REGION Network 14: EM - UnSuspending State Complete
   RUNG wire#powerrail
      Contact( "EM01".PackML_Sts.Alarm.sts_UnSuspending_SC )
      wire#w1
      Contact( "EM01".PackML_Sts.CM01.sts_UnSuspending_SC )
      wire#w2
      Contact( "EM01".PackML_Sts.CM02.sts_UnSuspending_SC )
      wire#w3
      Contact( "EM01".PackML_Sts.CM03.sts_UnSuspending_SC )
      wire#w4
      Contact( "EM01".PackML_Sts.CM04.sts_UnSuspending_SC )
      wire#w5
      Contact( "EM01".PackML_Sts.CM05.sts_UnSuspending_SC )
      wire#w6
      Contact( "EM01".PackML_Sts.CM06.sts_UnSuspending_SC )
      wire#w7
      Contact( "EM01".PackML_Sts.CM07.sts_UnSuspending_SC )
      wire#w8
      Contact( "EM01".PackML_Sts.CM08.sts_UnSuspending_SC )
      wire#w9
      Contact( "EM01".PackML_Sts.CM09.sts_UnSuspending_SC )
      wire#w10
      Contact( "EM01".PackML_Sts.CM10.sts_UnSuspending_SC )
      wire#w11
      Coil( "EM01".PackML_Sts.Unit.sts_UnSuspending_SC )
   END_RUNG
   RUNG wire#powerrail
      I_Contact( "EM01".PackML_Sts.Alarm.moduleActive )
   END_RUNG wire#w1
   RUNG wire#w1
      I_Contact( "EM01".PackML_Sts.CM01.moduleActive )
   END_RUNG wire#w2
   RUNG wire#w2
      I_Contact( "EM01".PackML_Sts.CM02.moduleActive )
   END_RUNG wire#w3
   RUNG wire#w3
      I_Contact( "EM01".PackML_Sts.CM03.moduleActive )
   END_RUNG wire#w4
   RUNG wire#w4
      I_Contact( "EM01".PackML_Sts.CM04.moduleActive )
   END_RUNG wire#w5
   RUNG wire#w5
      I_Contact( "EM01".PackML_Sts.CM05.moduleActive )
   END_RUNG wire#w6
   RUNG wire#w6
      I_Contact( "EM01".PackML_Sts.CM06.moduleActive )
   END_RUNG wire#w7
   RUNG wire#w7
      I_Contact( "EM01".PackML_Sts.CM07.moduleActive )
   END_RUNG wire#w8
   RUNG wire#w8
      I_Contact( "EM01".PackML_Sts.CM08.moduleActive )
   END_RUNG wire#w9
   RUNG wire#w9
      I_Contact( "EM01".PackML_Sts.CM09.moduleActive )
   END_RUNG wire#w10
   RUNG wire#w10
      I_Contact( "EM01".PackML_Sts.CM10.moduleActive )
   END_RUNG wire#w11
   // the same network as SCL:
   "EM01".PackML_Sts.Unit.sts_UnSuspending_SC := ("EM01".PackML_Sts.Alarm.sts_UnSuspending_SC OR NOT "EM01".PackML_Sts.Alarm.moduleActive) AND ("EM01".PackML_Sts.CM01.sts_UnSuspending_SC OR NOT "EM01".PackML_Sts.CM01.moduleActive) AND ("EM01".PackML_Sts.CM02.sts_UnSuspending_SC OR NOT "EM01".PackML_Sts.CM02.moduleActive) AND ("EM01".PackML_Sts.CM03.sts_UnSuspending_SC OR NOT "EM01".PackML_Sts.CM03.moduleActive) AND ("EM01".PackML_Sts.CM04.sts_UnSuspending_SC OR NOT "EM01".PackML_Sts.CM04.moduleActive) AND ("EM01".PackML_Sts.CM05.sts_UnSuspending_SC OR NOT "EM01".PackML_Sts.CM05.moduleActive) AND ("EM01".PackML_Sts.CM06.sts_UnSuspending_SC OR NOT "EM01".PackML_Sts.CM06.moduleActive) AND ("EM01".PackML_Sts.CM07.sts_UnSuspending_SC OR NOT "EM01".PackML_Sts.CM07.moduleActive) AND ("EM01".PackML_Sts.CM08.sts_UnSuspending_SC OR NOT "EM01".PackML_Sts.CM08.moduleActive) AND ("EM01".PackML_Sts.CM09.sts_UnSuspending_SC OR NOT "EM01".PackML_Sts.CM09.moduleActive) AND ("EM01".PackML_Sts.CM10.sts_UnSuspending_SC OR NOT "EM01".PackML_Sts.CM10.moduleActive);
END_REGION

REGION Network 15: EM - Abort Command
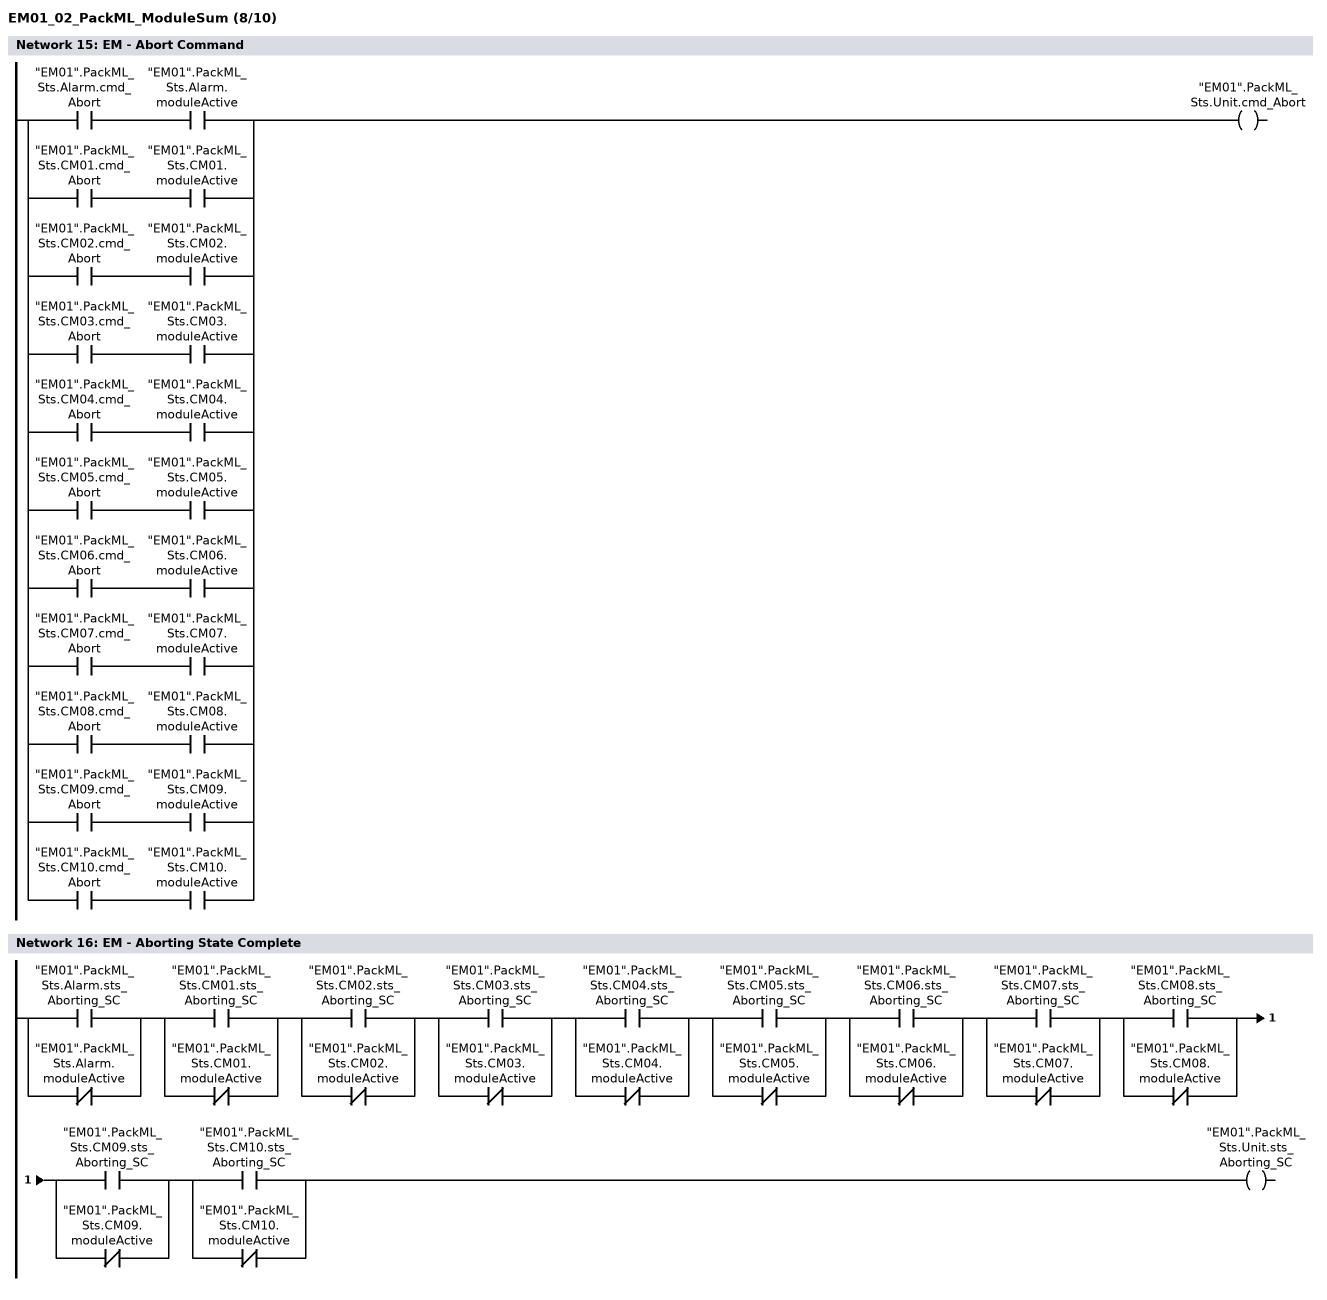
   RUNG wire#powerrail
      Contact( "EM01".PackML_Sts.Alarm.cmd_Abort )
      Contact( "EM01".PackML_Sts.Alarm.moduleActive )
      wire#w1
      Coil( "EM01".PackML_Sts.Unit.cmd_Abort )
   END_RUNG
   RUNG wire#powerrail
      Contact( "EM01".PackML_Sts.CM01.cmd_Abort )
      Contact( "EM01".PackML_Sts.CM01.moduleActive )
   END_RUNG wire#w1
   RUNG wire#powerrail
      Contact( "EM01".PackML_Sts.CM02.cmd_Abort )
      Contact( "EM01".PackML_Sts.CM02.moduleActive )
   END_RUNG wire#w1
   RUNG wire#powerrail
      Contact( "EM01".PackML_Sts.CM03.cmd_Abort )
      Contact( "EM01".PackML_Sts.CM03.moduleActive )
   END_RUNG wire#w1
   RUNG wire#powerrail
      Contact( "EM01".PackML_Sts.CM04.cmd_Abort )
      Contact( "EM01".PackML_Sts.CM04.moduleActive )
   END_RUNG wire#w1
   RUNG wire#powerrail
      Contact( "EM01".PackML_Sts.CM05.cmd_Abort )
      Contact( "EM01".PackML_Sts.CM05.moduleActive )
   END_RUNG wire#w1
   RUNG wire#powerrail
      Contact( "EM01".PackML_Sts.CM06.cmd_Abort )
      Contact( "EM01".PackML_Sts.CM06.moduleActive )
   END_RUNG wire#w1
   RUNG wire#powerrail
      Contact( "EM01".PackML_Sts.CM07.cmd_Abort )
      Contact( "EM01".PackML_Sts.CM07.moduleActive )
   END_RUNG wire#w1
   RUNG wire#powerrail
      Contact( "EM01".PackML_Sts.CM08.cmd_Abort )
      Contact( "EM01".PackML_Sts.CM08.moduleActive )
   END_RUNG wire#w1
   RUNG wire#powerrail
      Contact( "EM01".PackML_Sts.CM09.cmd_Abort )
      Contact( "EM01".PackML_Sts.CM09.moduleActive )
   END_RUNG wire#w1
   RUNG wire#powerrail
      Contact( "EM01".PackML_Sts.CM10.cmd_Abort )
      Contact( "EM01".PackML_Sts.CM10.moduleActive )
   END_RUNG wire#w1
   // the same network as SCL:
   "EM01".PackML_Sts.Unit.cmd_Abort := ("EM01".PackML_Sts.Alarm.cmd_Abort AND "EM01".PackML_Sts.Alarm.moduleActive) OR ("EM01".PackML_Sts.CM01.cmd_Abort AND "EM01".PackML_Sts.CM01.moduleActive) OR ("EM01".PackML_Sts.CM02.cmd_Abort AND "EM01".PackML_Sts.CM02.moduleActive) OR ("EM01".PackML_Sts.CM03.cmd_Abort AND "EM01".PackML_Sts.CM03.moduleActive) OR ("EM01".PackML_Sts.CM04.cmd_Abort AND "EM01".PackML_Sts.CM04.moduleActive) OR ("EM01".PackML_Sts.CM05.cmd_Abort AND "EM01".PackML_Sts.CM05.moduleActive) OR ("EM01".PackML_Sts.CM06.cmd_Abort AND "EM01".PackML_Sts.CM06.moduleActive) OR ("EM01".PackML_Sts.CM07.cmd_Abort AND "EM01".PackML_Sts.CM07.moduleActive) OR ("EM01".PackML_Sts.CM08.cmd_Abort AND "EM01".PackML_Sts.CM08.moduleActive) OR ("EM01".PackML_Sts.CM09.cmd_Abort AND "EM01".PackML_Sts.CM09.moduleActive) OR ("EM01".PackML_Sts.CM10.cmd_Abort AND "EM01".PackML_Sts.CM10.moduleActive);
END_REGION

REGION Network 16: EM - Aborting State Complete
   RUNG wire#powerrail
      Contact( "EM01".PackML_Sts.Alarm.sts_Aborting_SC )
      wire#w1
      Contact( "EM01".PackML_Sts.CM01.sts_Aborting_SC )
      wire#w2
      Contact( "EM01".PackML_Sts.CM02.sts_Aborting_SC )
      wire#w3
      Contact( "EM01".PackML_Sts.CM03.sts_Aborting_SC )
      wire#w4
      Contact( "EM01".PackML_Sts.CM04.sts_Aborting_SC )
      wire#w5
      Contact( "EM01".PackML_Sts.CM05.sts_Aborting_SC )
      wire#w6
      Contact( "EM01".PackML_Sts.CM06.sts_Aborting_SC )
      wire#w7
      Contact( "EM01".PackML_Sts.CM07.sts_Aborting_SC )
      wire#w8
      Contact( "EM01".PackML_Sts.CM08.sts_Aborting_SC )
      wire#w9
      Contact( "EM01".PackML_Sts.CM09.sts_Aborting_SC )
      wire#w10
      Contact( "EM01".PackML_Sts.CM10.sts_Aborting_SC )
      wire#w11
      Coil( "EM01".PackML_Sts.Unit.sts_Aborting_SC )
   END_RUNG
   RUNG wire#powerrail
      I_Contact( "EM01".PackML_Sts.Alarm.moduleActive )
   END_RUNG wire#w1
   RUNG wire#w1
      I_Contact( "EM01".PackML_Sts.CM01.moduleActive )
   END_RUNG wire#w2
   RUNG wire#w2
      I_Contact( "EM01".PackML_Sts.CM02.moduleActive )
   END_RUNG wire#w3
   RUNG wire#w3
      I_Contact( "EM01".PackML_Sts.CM03.moduleActive )
   END_RUNG wire#w4
   RUNG wire#w4
      I_Contact( "EM01".PackML_Sts.CM04.moduleActive )
   END_RUNG wire#w5
   RUNG wire#w5
      I_Contact( "EM01".PackML_Sts.CM05.moduleActive )
   END_RUNG wire#w6
   RUNG wire#w6
      I_Contact( "EM01".PackML_Sts.CM06.moduleActive )
   END_RUNG wire#w7
   RUNG wire#w7
      I_Contact( "EM01".PackML_Sts.CM07.moduleActive )
   END_RUNG wire#w8
   RUNG wire#w8
      I_Contact( "EM01".PackML_Sts.CM08.moduleActive )
   END_RUNG wire#w9
   RUNG wire#w9
      I_Contact( "EM01".PackML_Sts.CM09.moduleActive )
   END_RUNG wire#w10
   RUNG wire#w10
      I_Contact( "EM01".PackML_Sts.CM10.moduleActive )
   END_RUNG wire#w11
   // the same network as SCL:
   "EM01".PackML_Sts.Unit.sts_Aborting_SC := ("EM01".PackML_Sts.Alarm.sts_Aborting_SC OR NOT "EM01".PackML_Sts.Alarm.moduleActive) AND ("EM01".PackML_Sts.CM01.sts_Aborting_SC OR NOT "EM01".PackML_Sts.CM01.moduleActive) AND ("EM01".PackML_Sts.CM02.sts_Aborting_SC OR NOT "EM01".PackML_Sts.CM02.moduleActive) AND ("EM01".PackML_Sts.CM03.sts_Aborting_SC OR NOT "EM01".PackML_Sts.CM03.moduleActive) AND ("EM01".PackML_Sts.CM04.sts_Aborting_SC OR NOT "EM01".PackML_Sts.CM04.moduleActive) AND ("EM01".PackML_Sts.CM05.sts_Aborting_SC OR NOT "EM01".PackML_Sts.CM05.moduleActive) AND ("EM01".PackML_Sts.CM06.sts_Aborting_SC OR NOT "EM01".PackML_Sts.CM06.moduleActive) AND ("EM01".PackML_Sts.CM07.sts_Aborting_SC OR NOT "EM01".PackML_Sts.CM07.moduleActive) AND ("EM01".PackML_Sts.CM08.sts_Aborting_SC OR NOT "EM01".PackML_Sts.CM08.moduleActive) AND ("EM01".PackML_Sts.CM09.sts_Aborting_SC OR NOT "EM01".PackML_Sts.CM09.moduleActive) AND ("EM01".PackML_Sts.CM10.sts_Aborting_SC OR NOT "EM01".PackML_Sts.CM10.moduleActive);
END_REGION

REGION Network 17: EM - Clear Command
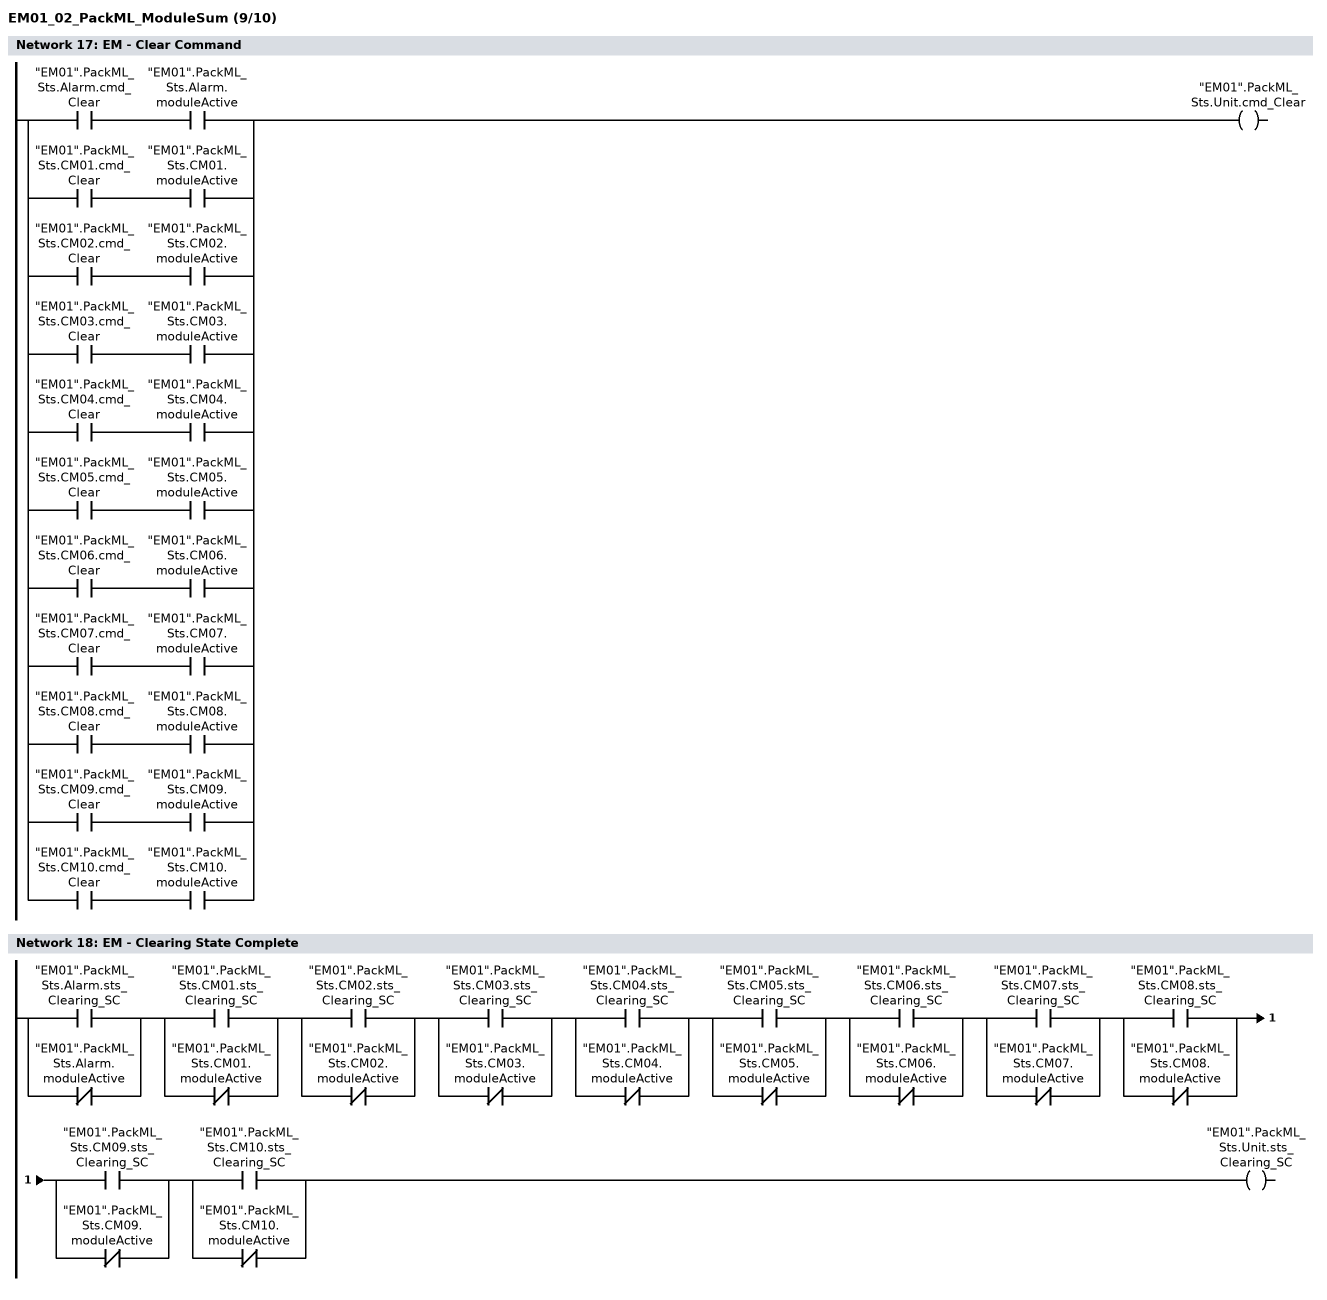
   RUNG wire#powerrail
      Contact( "EM01".PackML_Sts.Alarm.cmd_Clear )
      Contact( "EM01".PackML_Sts.Alarm.moduleActive )
      wire#w1
      Coil( "EM01".PackML_Sts.Unit.cmd_Clear )
   END_RUNG
   RUNG wire#powerrail
      Contact( "EM01".PackML_Sts.CM01.cmd_Clear )
      Contact( "EM01".PackML_Sts.CM01.moduleActive )
   END_RUNG wire#w1
   RUNG wire#powerrail
      Contact( "EM01".PackML_Sts.CM02.cmd_Clear )
      Contact( "EM01".PackML_Sts.CM02.moduleActive )
   END_RUNG wire#w1
   RUNG wire#powerrail
      Contact( "EM01".PackML_Sts.CM03.cmd_Clear )
      Contact( "EM01".PackML_Sts.CM03.moduleActive )
   END_RUNG wire#w1
   RUNG wire#powerrail
      Contact( "EM01".PackML_Sts.CM04.cmd_Clear )
      Contact( "EM01".PackML_Sts.CM04.moduleActive )
   END_RUNG wire#w1
   RUNG wire#powerrail
      Contact( "EM01".PackML_Sts.CM05.cmd_Clear )
      Contact( "EM01".PackML_Sts.CM05.moduleActive )
   END_RUNG wire#w1
   RUNG wire#powerrail
      Contact( "EM01".PackML_Sts.CM06.cmd_Clear )
      Contact( "EM01".PackML_Sts.CM06.moduleActive )
   END_RUNG wire#w1
   RUNG wire#powerrail
      Contact( "EM01".PackML_Sts.CM07.cmd_Clear )
      Contact( "EM01".PackML_Sts.CM07.moduleActive )
   END_RUNG wire#w1
   RUNG wire#powerrail
      Contact( "EM01".PackML_Sts.CM08.cmd_Clear )
      Contact( "EM01".PackML_Sts.CM08.moduleActive )
   END_RUNG wire#w1
   RUNG wire#powerrail
      Contact( "EM01".PackML_Sts.CM09.cmd_Clear )
      Contact( "EM01".PackML_Sts.CM09.moduleActive )
   END_RUNG wire#w1
   RUNG wire#powerrail
      Contact( "EM01".PackML_Sts.CM10.cmd_Clear )
      Contact( "EM01".PackML_Sts.CM10.moduleActive )
   END_RUNG wire#w1
   // the same network as SCL:
   "EM01".PackML_Sts.Unit.cmd_Clear := ("EM01".PackML_Sts.Alarm.cmd_Clear AND "EM01".PackML_Sts.Alarm.moduleActive) OR ("EM01".PackML_Sts.CM01.cmd_Clear AND "EM01".PackML_Sts.CM01.moduleActive) OR ("EM01".PackML_Sts.CM02.cmd_Clear AND "EM01".PackML_Sts.CM02.moduleActive) OR ("EM01".PackML_Sts.CM03.cmd_Clear AND "EM01".PackML_Sts.CM03.moduleActive) OR ("EM01".PackML_Sts.CM04.cmd_Clear AND "EM01".PackML_Sts.CM04.moduleActive) OR ("EM01".PackML_Sts.CM05.cmd_Clear AND "EM01".PackML_Sts.CM05.moduleActive) OR ("EM01".PackML_Sts.CM06.cmd_Clear AND "EM01".PackML_Sts.CM06.moduleActive) OR ("EM01".PackML_Sts.CM07.cmd_Clear AND "EM01".PackML_Sts.CM07.moduleActive) OR ("EM01".PackML_Sts.CM08.cmd_Clear AND "EM01".PackML_Sts.CM08.moduleActive) OR ("EM01".PackML_Sts.CM09.cmd_Clear AND "EM01".PackML_Sts.CM09.moduleActive) OR ("EM01".PackML_Sts.CM10.cmd_Clear AND "EM01".PackML_Sts.CM10.moduleActive);
END_REGION

REGION Network 18: EM - Clearing State Complete
   RUNG wire#powerrail
      Contact( "EM01".PackML_Sts.Alarm.sts_Clearing_SC )
      wire#w1
      Contact( "EM01".PackML_Sts.CM01.sts_Clearing_SC )
      wire#w2
      Contact( "EM01".PackML_Sts.CM02.sts_Clearing_SC )
      wire#w3
      Contact( "EM01".PackML_Sts.CM03.sts_Clearing_SC )
      wire#w4
      Contact( "EM01".PackML_Sts.CM04.sts_Clearing_SC )
      wire#w5
      Contact( "EM01".PackML_Sts.CM05.sts_Clearing_SC )
      wire#w6
      Contact( "EM01".PackML_Sts.CM06.sts_Clearing_SC )
      wire#w7
      Contact( "EM01".PackML_Sts.CM07.sts_Clearing_SC )
      wire#w8
      Contact( "EM01".PackML_Sts.CM08.sts_Clearing_SC )
      wire#w9
      Contact( "EM01".PackML_Sts.CM09.sts_Clearing_SC )
      wire#w10
      Contact( "EM01".PackML_Sts.CM10.sts_Clearing_SC )
      wire#w11
      Coil( "EM01".PackML_Sts.Unit.sts_Clearing_SC )
   END_RUNG
   RUNG wire#powerrail
      I_Contact( "EM01".PackML_Sts.Alarm.moduleActive )
   END_RUNG wire#w1
   RUNG wire#w1
      I_Contact( "EM01".PackML_Sts.CM01.moduleActive )
   END_RUNG wire#w2
   RUNG wire#w2
      I_Contact( "EM01".PackML_Sts.CM02.moduleActive )
   END_RUNG wire#w3
   RUNG wire#w3
      I_Contact( "EM01".PackML_Sts.CM03.moduleActive )
   END_RUNG wire#w4
   RUNG wire#w4
      I_Contact( "EM01".PackML_Sts.CM04.moduleActive )
   END_RUNG wire#w5
   RUNG wire#w5
      I_Contact( "EM01".PackML_Sts.CM05.moduleActive )
   END_RUNG wire#w6
   RUNG wire#w6
      I_Contact( "EM01".PackML_Sts.CM06.moduleActive )
   END_RUNG wire#w7
   RUNG wire#w7
      I_Contact( "EM01".PackML_Sts.CM07.moduleActive )
   END_RUNG wire#w8
   RUNG wire#w8
      I_Contact( "EM01".PackML_Sts.CM08.moduleActive )
   END_RUNG wire#w9
   RUNG wire#w9
      I_Contact( "EM01".PackML_Sts.CM09.moduleActive )
   END_RUNG wire#w10
   RUNG wire#w10
      I_Contact( "EM01".PackML_Sts.CM10.moduleActive )
   END_RUNG wire#w11
   // the same network as SCL:
   "EM01".PackML_Sts.Unit.sts_Clearing_SC := ("EM01".PackML_Sts.Alarm.sts_Clearing_SC OR NOT "EM01".PackML_Sts.Alarm.moduleActive) AND ("EM01".PackML_Sts.CM01.sts_Clearing_SC OR NOT "EM01".PackML_Sts.CM01.moduleActive) AND ("EM01".PackML_Sts.CM02.sts_Clearing_SC OR NOT "EM01".PackML_Sts.CM02.moduleActive) AND ("EM01".PackML_Sts.CM03.sts_Clearing_SC OR NOT "EM01".PackML_Sts.CM03.moduleActive) AND ("EM01".PackML_Sts.CM04.sts_Clearing_SC OR NOT "EM01".PackML_Sts.CM04.moduleActive) AND ("EM01".PackML_Sts.CM05.sts_Clearing_SC OR NOT "EM01".PackML_Sts.CM05.moduleActive) AND ("EM01".PackML_Sts.CM06.sts_Clearing_SC OR NOT "EM01".PackML_Sts.CM06.moduleActive) AND ("EM01".PackML_Sts.CM07.sts_Clearing_SC OR NOT "EM01".PackML_Sts.CM07.moduleActive) AND ("EM01".PackML_Sts.CM08.sts_Clearing_SC OR NOT "EM01".PackML_Sts.CM08.moduleActive) AND ("EM01".PackML_Sts.CM09.sts_Clearing_SC OR NOT "EM01".PackML_Sts.CM09.moduleActive) AND ("EM01".PackML_Sts.CM10.sts_Clearing_SC OR NOT "EM01".PackML_Sts.CM10.moduleActive);
END_REGION

REGION Network 19: EM - Execute State Complete
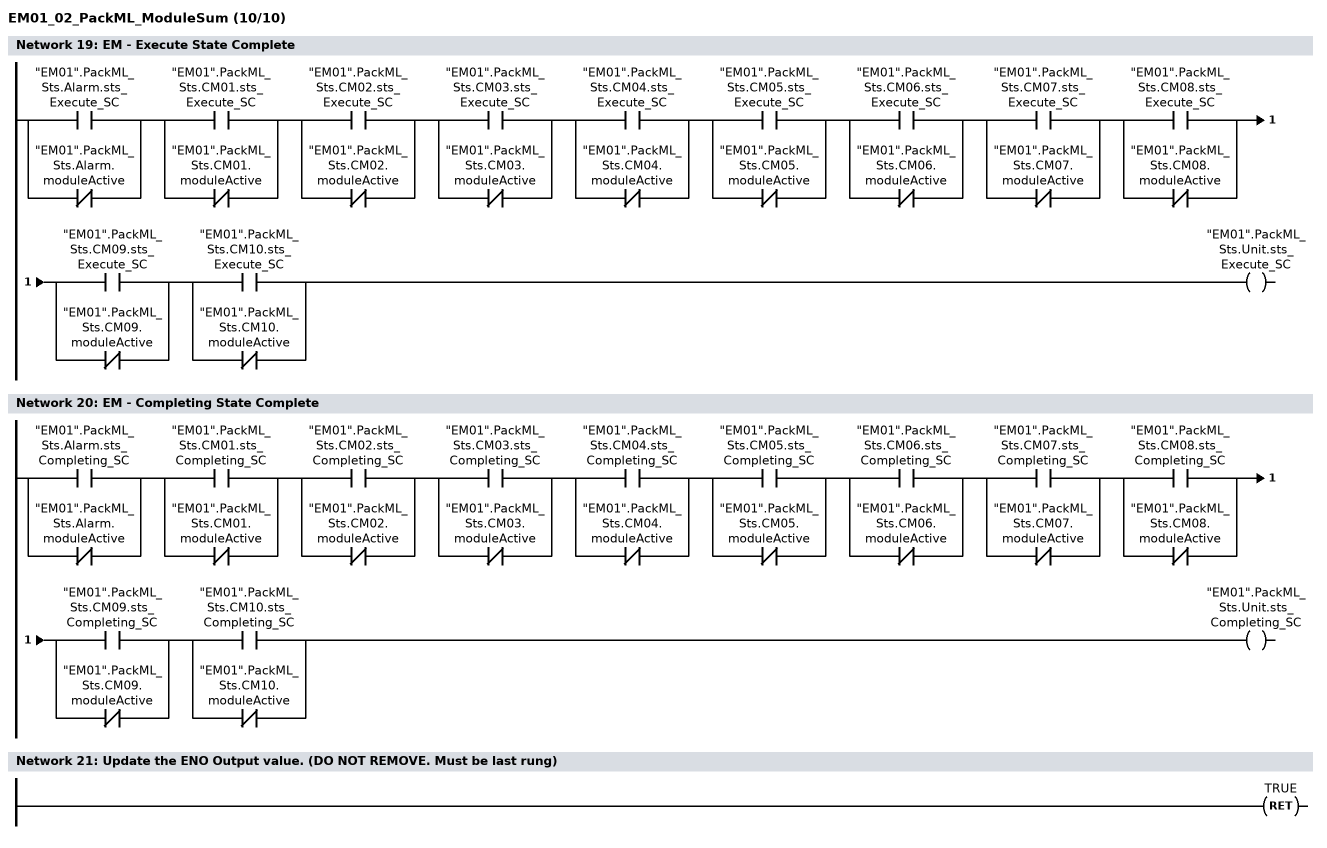
   RUNG wire#powerrail
      Contact( "EM01".PackML_Sts.Alarm.sts_Execute_SC )
      wire#w1
      Contact( "EM01".PackML_Sts.CM01.sts_Execute_SC )
      wire#w2
      Contact( "EM01".PackML_Sts.CM02.sts_Execute_SC )
      wire#w3
      Contact( "EM01".PackML_Sts.CM03.sts_Execute_SC )
      wire#w4
      Contact( "EM01".PackML_Sts.CM04.sts_Execute_SC )
      wire#w5
      Contact( "EM01".PackML_Sts.CM05.sts_Execute_SC )
      wire#w6
      Contact( "EM01".PackML_Sts.CM06.sts_Execute_SC )
      wire#w7
      Contact( "EM01".PackML_Sts.CM07.sts_Execute_SC )
      wire#w8
      Contact( "EM01".PackML_Sts.CM08.sts_Execute_SC )
      wire#w9
      Contact( "EM01".PackML_Sts.CM09.sts_Execute_SC )
      wire#w10
      Contact( "EM01".PackML_Sts.CM10.sts_Execute_SC )
      wire#w11
      Coil( "EM01".PackML_Sts.Unit.sts_Execute_SC )
   END_RUNG
   RUNG wire#powerrail
      I_Contact( "EM01".PackML_Sts.Alarm.moduleActive )
   END_RUNG wire#w1
   RUNG wire#w1
      I_Contact( "EM01".PackML_Sts.CM01.moduleActive )
   END_RUNG wire#w2
   RUNG wire#w2
      I_Contact( "EM01".PackML_Sts.CM02.moduleActive )
   END_RUNG wire#w3
   RUNG wire#w3
      I_Contact( "EM01".PackML_Sts.CM03.moduleActive )
   END_RUNG wire#w4
   RUNG wire#w4
      I_Contact( "EM01".PackML_Sts.CM04.moduleActive )
   END_RUNG wire#w5
   RUNG wire#w5
      I_Contact( "EM01".PackML_Sts.CM05.moduleActive )
   END_RUNG wire#w6
   RUNG wire#w6
      I_Contact( "EM01".PackML_Sts.CM06.moduleActive )
   END_RUNG wire#w7
   RUNG wire#w7
      I_Contact( "EM01".PackML_Sts.CM07.moduleActive )
   END_RUNG wire#w8
   RUNG wire#w8
      I_Contact( "EM01".PackML_Sts.CM08.moduleActive )
   END_RUNG wire#w9
   RUNG wire#w9
      I_Contact( "EM01".PackML_Sts.CM09.moduleActive )
   END_RUNG wire#w10
   RUNG wire#w10
      I_Contact( "EM01".PackML_Sts.CM10.moduleActive )
   END_RUNG wire#w11
   // the same network as SCL:
   "EM01".PackML_Sts.Unit.sts_Execute_SC := ("EM01".PackML_Sts.Alarm.sts_Execute_SC OR NOT "EM01".PackML_Sts.Alarm.moduleActive) AND ("EM01".PackML_Sts.CM01.sts_Execute_SC OR NOT "EM01".PackML_Sts.CM01.moduleActive) AND ("EM01".PackML_Sts.CM02.sts_Execute_SC OR NOT "EM01".PackML_Sts.CM02.moduleActive) AND ("EM01".PackML_Sts.CM03.sts_Execute_SC OR NOT "EM01".PackML_Sts.CM03.moduleActive) AND ("EM01".PackML_Sts.CM04.sts_Execute_SC OR NOT "EM01".PackML_Sts.CM04.moduleActive) AND ("EM01".PackML_Sts.CM05.sts_Execute_SC OR NOT "EM01".PackML_Sts.CM05.moduleActive) AND ("EM01".PackML_Sts.CM06.sts_Execute_SC OR NOT "EM01".PackML_Sts.CM06.moduleActive) AND ("EM01".PackML_Sts.CM07.sts_Execute_SC OR NOT "EM01".PackML_Sts.CM07.moduleActive) AND ("EM01".PackML_Sts.CM08.sts_Execute_SC OR NOT "EM01".PackML_Sts.CM08.moduleActive) AND ("EM01".PackML_Sts.CM09.sts_Execute_SC OR NOT "EM01".PackML_Sts.CM09.moduleActive) AND ("EM01".PackML_Sts.CM10.sts_Execute_SC OR NOT "EM01".PackML_Sts.CM10.moduleActive);
END_REGION

REGION Network 20: EM - Completing State Complete
   RUNG wire#powerrail
      Contact( "EM01".PackML_Sts.Alarm.sts_Completing_SC )
      wire#w1
      Contact( "EM01".PackML_Sts.CM01.sts_Completing_SC )
      wire#w2
      Contact( "EM01".PackML_Sts.CM02.sts_Completing_SC )
      wire#w3
      Contact( "EM01".PackML_Sts.CM03.sts_Completing_SC )
      wire#w4
      Contact( "EM01".PackML_Sts.CM04.sts_Completing_SC )
      wire#w5
      Contact( "EM01".PackML_Sts.CM05.sts_Completing_SC )
      wire#w6
      Contact( "EM01".PackML_Sts.CM06.sts_Completing_SC )
      wire#w7
      Contact( "EM01".PackML_Sts.CM07.sts_Completing_SC )
      wire#w8
      Contact( "EM01".PackML_Sts.CM08.sts_Completing_SC )
      wire#w9
      Contact( "EM01".PackML_Sts.CM09.sts_Completing_SC )
      wire#w10
      Contact( "EM01".PackML_Sts.CM10.sts_Completing_SC )
      wire#w11
      Coil( "EM01".PackML_Sts.Unit.sts_Completing_SC )
   END_RUNG
   RUNG wire#powerrail
      I_Contact( "EM01".PackML_Sts.Alarm.moduleActive )
   END_RUNG wire#w1
   RUNG wire#w1
      I_Contact( "EM01".PackML_Sts.CM01.moduleActive )
   END_RUNG wire#w2
   RUNG wire#w2
      I_Contact( "EM01".PackML_Sts.CM02.moduleActive )
   END_RUNG wire#w3
   RUNG wire#w3
      I_Contact( "EM01".PackML_Sts.CM03.moduleActive )
   END_RUNG wire#w4
   RUNG wire#w4
      I_Contact( "EM01".PackML_Sts.CM04.moduleActive )
   END_RUNG wire#w5
   RUNG wire#w5
      I_Contact( "EM01".PackML_Sts.CM05.moduleActive )
   END_RUNG wire#w6
   RUNG wire#w6
      I_Contact( "EM01".PackML_Sts.CM06.moduleActive )
   END_RUNG wire#w7
   RUNG wire#w7
      I_Contact( "EM01".PackML_Sts.CM07.moduleActive )
   END_RUNG wire#w8
   RUNG wire#w8
      I_Contact( "EM01".PackML_Sts.CM08.moduleActive )
   END_RUNG wire#w9
   RUNG wire#w9
      I_Contact( "EM01".PackML_Sts.CM09.moduleActive )
   END_RUNG wire#w10
   RUNG wire#w10
      I_Contact( "EM01".PackML_Sts.CM10.moduleActive )
   END_RUNG wire#w11
   // the same network as SCL:
   "EM01".PackML_Sts.Unit.sts_Completing_SC := ("EM01".PackML_Sts.Alarm.sts_Completing_SC OR NOT "EM01".PackML_Sts.Alarm.moduleActive) AND ("EM01".PackML_Sts.CM01.sts_Completing_SC OR NOT "EM01".PackML_Sts.CM01.moduleActive) AND ("EM01".PackML_Sts.CM02.sts_Completing_SC OR NOT "EM01".PackML_Sts.CM02.moduleActive) AND ("EM01".PackML_Sts.CM03.sts_Completing_SC OR NOT "EM01".PackML_Sts.CM03.moduleActive) AND ("EM01".PackML_Sts.CM04.sts_Completing_SC OR NOT "EM01".PackML_Sts.CM04.moduleActive) AND ("EM01".PackML_Sts.CM05.sts_Completing_SC OR NOT "EM01".PackML_Sts.CM05.moduleActive) AND ("EM01".PackML_Sts.CM06.sts_Completing_SC OR NOT "EM01".PackML_Sts.CM06.moduleActive) AND ("EM01".PackML_Sts.CM07.sts_Completing_SC OR NOT "EM01".PackML_Sts.CM07.moduleActive) AND ("EM01".PackML_Sts.CM08.sts_Completing_SC OR NOT "EM01".PackML_Sts.CM08.moduleActive) AND ("EM01".PackML_Sts.CM09.sts_Completing_SC OR NOT "EM01".PackML_Sts.CM09.moduleActive) AND ("EM01".PackML_Sts.CM10.sts_Completing_SC OR NOT "EM01".PackML_Sts.CM10.moduleActive);
END_REGION

REGION Network 21: Update the ENO Output value. (DO NOT REMOVE. Must be last rung)
   RUNG wire#powerrail
      ReturnCoil( TRUE )
   END_RUNG
   // the same network as SCL:
   ENO := TRUE;
   RETURN;
END_REGION
END_FUNCTION_BLOCK

FUNCTION_BLOCK "EM01_CM01_Conveyor"   // FB31671, LAD
TITLE = EM01_CM01
{ S7_Optimized_Access := 'TRUE' }
AUTHOR : tech.team.motioncontrol@siemens.com
FAMILY : CPG
VERSION : 1.1
// Support: tech.team.motioncontrol@siemens.com
   VAR
      statDummyBool : Bool;   // dummy bool - placeholder
      instBeltConveyor : "BeltConveyor";
   END_VAR
BEGIN

REGION Network 1: *** Begin the Setpoint Management Information Section ***
END_REGION

REGION Network 2: *** Begin the Logic Section ***
END_REGION

REGION Network 3: Belt conveyor instance
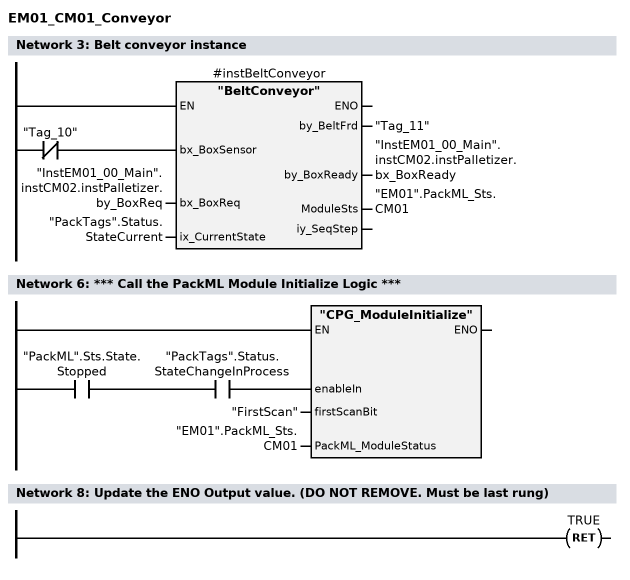
   RUNG wire#powerrail
      #instBeltConveyor(bx_BoxSensor := wire#w1, bx_BoxReq := "InstEM01_00_Main".instCM02.instPalletizer.by_BoxReq, ix_CurrentState := "PackTags".Status.StateCurrent, by_BeltFrd => "Tag_11", by_BoxReady => "InstEM01_00_Main".instCM02.instPalletizer.bx_BoxReady, ModuleSts => "EM01".PackML_Sts.CM01, iy_SeqStep =>)
   END_RUNG
   RUNG wire#powerrail
      I_Contact( "Tag_10" )
   END_RUNG wire#w1
   // the same network as SCL:
   #instBeltConveyor(bx_BoxSensor := NOT "Tag_10",   // "BeltConveyor"
                     bx_BoxReq := "InstEM01_00_Main".instCM02.instPalletizer.by_BoxReq,
                     ix_CurrentState := "PackTags".Status.StateCurrent,
                     by_BeltFrd => "Tag_11",
                     by_BoxReady => "InstEM01_00_Main".instCM02.instPalletizer.bx_BoxReady,
                     ModuleSts => "EM01".PackML_Sts.CM01);
END_REGION

REGION Network 4: *** Begin the Event Information Section ***
END_REGION

REGION Network 5: *** Begin the State Model Status Feedback Section ***
END_REGION

REGION Network 6: *** Call the PackML Module Initialize Logic ***
   RUNG wire#powerrail
      "CPG_ModuleInitialize"(enableIn := wire#w1, firstScanBit := "FirstScan", PackML_ModuleStatus := "EM01".PackML_Sts.CM01)
   END_RUNG
   RUNG wire#powerrail
      Contact( "PackML".Sts.State.Stopped )
      Contact( "PackTags".Status.StateChangeInProcess )
   END_RUNG wire#w1
   // the same network as SCL:
   "CPG_ModuleInitialize"(enableIn := "PackML".Sts.State.Stopped AND "PackTags".Status.StateChangeInProcess,
                          firstScanBit := "FirstScan",
                          PackML_ModuleStatus := "EM01".PackML_Sts.CM01);
END_REGION

REGION Network 8: Update the ENO Output value. (DO NOT REMOVE. Must be last rung)
   RUNG wire#powerrail
      ReturnCoil( TRUE )
   END_RUNG
   // the same network as SCL:
   ENO := TRUE;
   RETURN;
END_REGION
END_FUNCTION_BLOCK

FUNCTION_BLOCK "EM01_CM02_Palletizer"   // FB31672, LAD
TITLE = EM01_CM02
{ S7_Optimized_Access := 'TRUE' }
AUTHOR : tech.team.motioncontrol@siemens.com
FAMILY : CPG
VERSION : 1.1
// Support: tech.team.motioncontrol@siemens.com
   VAR
      statDummyBool : Bool;   // dummy bool - placeholder
      instPalletizer : "Palletizer";
      Ntrig : Bool;
   END_VAR
   VAR_TEMP   // added for the SCL form of the ladder/FBD networks
      _w1 : Bool;
   END_VAR
BEGIN

REGION Network 1: *** Begin the Setpoint Management Information Section ***
END_REGION

REGION Network 2: *** Begin the Logic Section ***
END_REGION

REGION Network 3: Palletizer instance